VAR_GLOBAL   // PLC tag table "Carrier_SDC_TagTable"
   "Carrier_01_Status" AT %IW400 : Word;   // CARRIER STATUS WORD
   "Carrier_01_Status.0" AT %I400.0 : Bool;   // HEARTBEAT
   "Carrier_01_Status.1" AT %I400.1 : Bool;   // MANUAL
   "Carrier_01_Status.2" AT %I400.2 : Bool;   // IN_AUTO
   "Carrier_01_Status.3" AT %I400.3 : Bool;   // POSITIONING_COMPLETE
   "Carrier_01_Status.4" AT %I400.4 : Bool;   // PRODUCTION HOLD
   "Carrier_01_Status.5" AT %I400.5 : Bool;   // CARRIER MOVING FORWARD
   "Carrier_01_Status.6" AT %I400.6 : Bool;   // CARRIER MOVING REVERSE
   "Carrier_01_Status.7" AT %I400.7 : Bool;   // CARRIER FAULT
   "Carrier_01_Status.8" AT %I401.0 : Bool;   // CRASH DETECT TRIPPED
   "Carrier_01_Status.9" AT %I401.1 : Bool;
   "Carrier_01_Status.10" AT %I401.2 : Bool;
   "Carrier_01_Status.11" AT %I401.3 : Bool;
   "Carrier_01_Status.12" AT %I401.4 : Bool;
   "Carrier_01_Status.13" AT %I401.5 : Bool;
   "Carrier_01_Status.14" AT %I401.6 : Bool;
   "Carrier_01_Status.15" AT %I401.7 : Bool;
   "Carrier_01_SDCFaultCode" AT %IW402 : Word;   // SDC FAULT CODE
   "Carrier_01_CarrierPosition" AT %ID404 : DWord;   // CARRIER POSITION
   "Carrier_01_CarrierNumber" AT %IW408 : Word;   // CARRIER NUMBER
   "Carrier_01_G120DControlWord" AT %IW410 : Word;   // G120D_STW1_CONTROL
   "Carrier_01_G120DControlWord.0" AT %I410.0 : Bool;   // Bit_00_ON
   "Carrier_01_G120DControlWord.1" AT %I410.1 : Bool;   // Bit_01_AUS2_INH
   "Carrier_01_G120DControlWord.2" AT %I410.2 : Bool;   // Bit_02_AUS3_STOP
   "Carrier_01_G120DControlWord.3" AT %I410.3 : Bool;   // Bit_03_EN
   "Carrier_01_G120DControlWord.4" AT %I410.4 : Bool;   // Bit_04_EN_RAMP
   "Carrier_01_G120DControlWord.5" AT %I410.5 : Bool;   // Bit_05_START_RAMP
   "Carrier_01_G120DControlWord.6" AT %I410.6 : Bool;   // Bit_06_SETPOINT
   "Carrier_01_G120DControlWord.7" AT %I410.7 : Bool;   // Bit_07_RESET
   "Carrier_01_G120DControlWord.8" AT %I411.0 : Bool;   // Bit_08_JOG_R
   "Carrier_01_G120DControlWord.9" AT %I411.1 : Bool;   // Bit_09_JOG_L
   "Carrier_01_G120DControlWord.10" AT %I411.2 : Bool;   // Bit_10_CONTR_PLC
   "Carrier_01_G120DControlWord.11" AT %I411.3 : Bool;   // Bit_11_REVERSE
   "Carrier_01_G120DControlWord.12" AT %I411.4 : Bool;   // Bit_12_BRAKE_RELEASE
   "Carrier_01_G120DControlWord.13" AT %I411.5 : Bool;   // Bit_13_DDS
   "Carrier_01_G120DControlWord.14" AT %I411.6 : Bool;   // Bit_14_DO0
   "Carrier_01_G120DControlWord.15" AT %I411.7 : Bool;   // Bit_15_DO1
   "Carrier_01_G120DStatusWord" AT %IW412 : Word;   // G120D_ZSW1_STATUS
   "Carrier_01_G120DStatusWord.0" AT %I412.0 : Bool;   // Bit_00_READY_RUN
   "Carrier_01_G120DStatusWord.1" AT %I412.1 : Bool;   // Bit_01_READY_ON
   "Carrier_01_G120DStatusWord.2" AT %I412.2 : Bool;   // Bit_02_ENABLE
   "Carrier_01_G120DStatusWord.3" AT %I412.3 : Bool;   // Bit_03_FAULT
   "Carrier_01_G120DStatusWord.4" AT %I412.4 : Bool;   // Bit_04_OFF2
   "Carrier_01_G120DStatusWord.5" AT %I412.5 : Bool;   // Bit_05_OFF3
   "Carrier_01_G120DStatusWord.6" AT %I412.6 : Bool;   // Bit_06_LOCK_OUT
   "Carrier_01_G120DStatusWord.7" AT %I412.7 : Bool;   // Bit_07_WARN
   "Carrier_01_G120DStatusWord.8" AT %I413.0 : Bool;   // Bit_08_NO_DEVIATION
   "Carrier_01_G120DStatusWord.9" AT %I413.1 : Bool;   // Bit_09_CONTR_PLC
   "Carrier_01_G120DStatusWord.10" AT %I413.2 : Bool;   // Bit_10_F_MAX
   "Carrier_01_G120DStatusWord.11" AT %I413.3 : Bool;   // Bit_11_LIMIT_REACHED
   "Carrier_01_G120DStatusWord.12" AT %I413.4 : Bool;   // Bit_12_BRAKE_OPEN
   "Carrier_01_G120DStatusWord.13" AT %I413.5 : Bool;   // Bit_13_NO_OVERTEMP
   "Carrier_01_G120DStatusWord.14" AT %I413.6 : Bool;   // Bit_14_CW_CCW
   "Carrier_01_G120DStatusWord.15" AT %I413.7 : Bool;   // Bit_15_OVERL
   "Carrier_01_Slot2_Input" AT %IW414 : Word;   // SLOT 2 INPUT WORD
   "Carrier_01_CrashDetectSW" AT %I414.0 : Bool;   // CRASH DETECT SW
   "Carrier_01_SpareSafetyInput(2_1)" AT %I414.1 : Bool;   // SPARE SAFETY INPUT
   "Carrier_01_SpareSafetyInput(2_2)" AT %I414.2 : Bool;   // SPARE SAFETY INPUT
   "Carrier_01_SpareSafetyInput(2_3)" AT %I414.3 : Bool;   // SPARE SAFETY INPUT
   "Carrier_01_SpareSafetyInput(2_4)" AT %I414.4 : Bool;   // SPARE SAFETY INPUT
   "Carrier_01_SpareSafetyInput(2_5)" AT %I414.5 : Bool;   // SPARE SAFETY INPUT
   "Carrier_01_SpareSafetyInput(2_6)" AT %I414.6 : Bool;   // SPARE SAFETY INPUT
   "Carrier_01_SpareSafetyInput(2_7)" AT %I414.7 : Bool;   // SPARE SAFETY INPUT
   "Carrier_01_Slot3_SafetyOutput" AT %IW415 : Word;   // SLOT 3 SAFETY OUTPUT WORD
   "Carrier_01_Crash_Detect_OK" AT %I415.0 : Bool;   // CARRIER CRASH DETECT
   "Carrier_01_SpareSafetyOutput(3_1)" AT %I415.1 : Bool;   // SPARE SAFETY OUTPUT
   "Carrier_01_SpareSafetyOutput(3_2)" AT %I415.2 : Bool;   // SPARE SAFETY OUTPUT
   "Carrier_01_SpareSafetyOutput(3_3)" AT %I415.3 : Bool;   // SPARE SAFETY OUTPUT
   "Carrier_01_SpareSafetyOutput(3_4)" AT %I415.4 : Bool;   // SPARE SAFETY OUTPUT
   "Carrier_01_SpareSafetyOutput(3_5)" AT %I415.5 : Bool;   // SPARE SAFETY OUTPUT
   "Carrier_01_SpareSafetyOutput(3_6)" AT %I415.6 : Bool;   // SPARE SAFETY OUTPUT
   "Carrier_01_SpareSafetyOutput(3_7)" AT %I415.7 : Bool;   // SPARE SAFETY OUTPUT
   "Carrier_01_Slot4_Input" AT %IW416 : Word;   // SLOT 4 INPUT WORD
   "Carrier_01_480VPowerOn_MDCB1" AT %I416.0 : Bool;   // 480 VAC POWER ON MDCB 1
   "Carrier_01_SpareInput(4_1)" AT %I416.1 : Bool;   // SPARE INPUT
   "Carrier_01_SpareInput(4_2)" AT %I416.2 : Bool;   // SPARE INPUT
   "Carrier_01_SitopSelectStatus" AT %I416.3 : Bool;   // SITOP SELECT STATUS
   "Carrier_01_DCsupplyOnPSCB2" AT %I416.4 : Bool;   // DC SUPPLY ON PSCB 2
   "Carrier_01_SpareInput(4_5)" AT %I416.5 : Bool;   // SPARE INPUT
   "Carrier_01_SpareInput(4_6)" AT %I416.6 : Bool;   // SPARE INPUT
   "Carrier_01_SpareInput(4_7)" AT %I416.7 : Bool;   // SPARE INPUT
   "Carrier_01_PB1_ProdHoldLH" AT %I417.0 : Bool;   // PB 1 PRODUCTION HOLD LH
   "Carrier_01_PB2_ResetLH" AT %I417.1 : Bool;   // PB 2 RESET LH
   "Carrier_01_PB3_ProdHoldRH" AT %I417.2 : Bool;   // PB 3 PRODUCTION HOLD RH
   "Carrier_01_PB4_ResetRH" AT %I417.3 : Bool;   // PB 4 RESET RH
   "Carrier_01_SpareInput(4_14)" AT %I417.4 : Bool;   // SPARE INPUT
   "Carrier_01_SpareInput(4_15)" AT %I417.5 : Bool;   // SPARE INPUT
   "Carrier_01_SpareInput(4_16)" AT %I417.6 : Bool;   // SPARE INPUT
   "Carrier_01_SpareInput(4_17)" AT %I417.7 : Bool;   // SPARE INPUT
   "Carrier_01_Slot5_Output" AT %IW418 : Word;   // SLOT 5 OUTPUT WORD
   "Carrier_01_IRD400_HMI_24VDC_ENABLE" AT %I418.0 : Bool;   // IRD 400 PANEL HMI 24V DC POWER
   "Carrier_01_FaultLight_LH" AT %I418.1 : Bool;   // FAULT LIGHT LH
   "Carrier_01_RunLight_LH" AT %I418.2 : Bool;   // RUN LIGHT LH
   "Carrier_01_FaultLight_RH" AT %I418.3 : Bool;   // FAULT LIGHT RH
   "Carrier_01_RunLight_RH" AT %I418.4 : Bool;   // RUN LIGHT RH
   "Carrier_01_SpareOutput(5_5)" AT %I418.5 : Bool;   // SPARE OUTPUT
   "Carrier_01_SpareOutput(5_6)" AT %I418.6 : Bool;   // SPARE OUTPUT
   "Carrier_01_SpareOutput(5_7)" AT %I418.7 : Bool;   // SPARE OUTPUT
   "Carrier_01_ActualSpeed" AT %IW420 : Word;   // ACTUAL SPEED
   "Carrier_01_CarrierDriveAlarm" AT %IW422 : Word;   // CARRIER DRIVE ALARM
   "Carrier_01_CarrierDriveWarning" AT %IW424 : Word;   // CARRIER DRIVE WARNING
   "Carrier_02_Status" AT %IW450 : Word;   // CARRIER STATUS WORD
   "Carrier_02_Status.0" AT %I450.0 : Bool;   // HEARTBEAT
   "Carrier_02_Status.1" AT %I450.1 : Bool;   // MANUAL
   "Carrier_02_Status.2" AT %I450.2 : Bool;   // IN_AUTO
   "Carrier_02_Status.3" AT %I450.3 : Bool;   // POSITIONING_COMPLETE
   "Carrier_02_Status.4" AT %I450.4 : Bool;   // PRODUCTION HOLD
   "Carrier_02_Status.5" AT %I450.5 : Bool;   // CARRIER MOVING FORWARD
   "Carrier_02_Status.6" AT %I450.6 : Bool;   // CARRIER MOVING REVERSE
   "Carrier_02_Status.7" AT %I450.7 : Bool;   // CARRIER FAULT
   "Carrier_02_Status.8" AT %I451.0 : Bool;   // CRASH DETECT TRIPPED
   "Carrier_02_Status.9" AT %I451.1 : Bool;
   "Carrier_02_Status.10" AT %I451.2 : Bool;
   "Carrier_02_Status.11" AT %I451.3 : Bool;
   "Carrier_02_Status.12" AT %I451.4 : Bool;
   "Carrier_02_Status.13" AT %I451.5 : Bool;
   "Carrier_02_Status.14" AT %I451.6 : Bool;
   "Carrier_02_Status.15" AT %I451.7 : Bool;
   "Carrier_02_SDCFaultCode" AT %IW452 : Word;   // SDC FAULT CODE
   "Carrier_02_CarrierPosition" AT %ID454 : DWord;   // CARRIER POSITION
   "Carrier_02_CarrierNumber" AT %IW458 : Word;   // CARRIER NUMBER
   "Carrier_02_G120DControlWord" AT %IW460 : Word;   // G120D_STW1_CONTROL
   "Carrier_02_G120DControlWord.0" AT %I460.0 : Bool;   // Bit_00_ON
   "Carrier_02_G120DControlWord.1" AT %I460.1 : Bool;   // Bit_01_AUS2_INH
   "Carrier_02_G120DControlWord.2" AT %I460.2 : Bool;   // Bit_02_AUS3_STOP
   "Carrier_02_G120DControlWord.3" AT %I460.3 : Bool;   // Bit_03_EN
   "Carrier_02_G120DControlWord.4" AT %I460.4 : Bool;   // Bit_04_EN_RAMP
   "Carrier_02_G120DControlWord.5" AT %I460.5 : Bool;   // Bit_05_START_RAMP
   "Carrier_02_G120DControlWord.6" AT %I460.6 : Bool;   // Bit_06_SETPOINT
   "Carrier_02_G120DControlWord.7" AT %I460.7 : Bool;   // Bit_07_RESET
   "Carrier_02_G120DControlWord.8" AT %I461.0 : Bool;   // Bit_08_JOG_R
   "Carrier_02_G120DControlWord.9" AT %I461.1 : Bool;   // Bit_09_JOG_L
   "Carrier_02_G120DControlWord.10" AT %I461.2 : Bool;   // Bit_10_CONTR_PLC
   "Carrier_02_G120DControlWord.11" AT %I461.3 : Bool;   // Bit_11_REVERSE
   "Carrier_02_G120DControlWord.12" AT %I461.4 : Bool;   // Bit_12_BRAKE_RELEASE
   "Carrier_02_G120DControlWord.13" AT %I461.5 : Bool;   // Bit_13_DDS
   "Carrier_02_G120DControlWord.14" AT %I461.6 : Bool;   // Bit_14_DO0
   "Carrier_02_G120DControlWord.15" AT %I461.7 : Bool;   // Bit_15_DO1
   "Carrier_02_G120DStatusWord" AT %IW462 : Word;   // G120D_ZSW1_STATUS
   "Carrier_02_G120DStatusWord.0" AT %I462.0 : Bool;   // Bit_00_READY_RUN
   "Carrier_02_G120DStatusWord.1" AT %I462.1 : Bool;   // Bit_01_READY_ON
   "Carrier_02_G120DStatusWord.2" AT %I462.2 : Bool;   // Bit_02_ENABLE
   "Carrier_02_G120DStatusWord.3" AT %I462.3 : Bool;   // Bit_03_FAULT
   "Carrier_02_G120DStatusWord.4" AT %I462.4 : Bool;   // Bit_04_OFF2
   "Carrier_02_G120DStatusWord.5" AT %I462.5 : Bool;   // Bit_05_OFF3
   "Carrier_02_G120DStatusWord.6" AT %I462.6 : Bool;   // Bit_06_LOCK_OUT
   "Carrier_02_G120DStatusWord.7" AT %I462.7 : Bool;   // Bit_07_WARN
   "Carrier_02_G120DStatusWord.8" AT %I463.0 : Bool;   // Bit_08_NO_DEVIATION
   "Carrier_02_G120DStatusWord.9" AT %I463.1 : Bool;   // Bit_09_CONTR_PLC
   "Carrier_02_G120DStatusWord.10" AT %I463.2 : Bool;   // Bit_10_F_MAX
   "Carrier_02_G120DStatusWord.11" AT %I463.3 : Bool;   // Bit_11_LIMIT_REACHED
   "Carrier_02_G120DStatusWord.12" AT %I463.4 : Bool;   // Bit_12_BRAKE_OPEN
   "Carrier_02_G120DStatusWord.13" AT %I463.5 : Bool;   // Bit_13_NO_OVERTEMP
   "Carrier_02_G120DStatusWord.14" AT %I463.6 : Bool;   // Bit_14_CW_CCW
   "Carrier_02_G120DStatusWord.15" AT %I463.7 : Bool;   // Bit_15_OVERL
   "Carrier_02_Slot2_Input" AT %IW464 : Word;   // SLOT 2 INPUT WORD
   "Carrier_02_CrashDetectSW" AT %I464.0 : Bool;   // CRASH DETECT SW
   "Carrier_02_SpareSafetyInput(2_1)" AT %I464.1 : Bool;   // SPARE SAFETY INPUT
   "Carrier_02_SpareSafetyInput(2_2)" AT %I464.2 : Bool;   // SPARE SAFETY INPUT
   "Carrier_02_SpareSafetyInput(2_3)" AT %I464.3 : Bool;   // SPARE SAFETY INPUT
   "Carrier_02_SpareSafetyInput(2_4)" AT %I464.4 : Bool;   // SPARE SAFETY INPUT
   "Carrier_02_SpareSafetyInput(2_5)" AT %I464.5 : Bool;   // SPARE SAFETY INPUT
   "Carrier_02_SpareSafetyInput(2_6)" AT %I464.6 : Bool;   // SPARE SAFETY INPUT
   "Carrier_02_SpareSafetyInput(2_7)" AT %I464.7 : Bool;   // SPARE SAFETY INPUT
   "Carrier_02_Slot3_SafetyOutput" AT %IW465 : Word;   // SLOT 3 SAFETY OUTPUT WORD
   "Carrier_02_Crash_Detect_OK" AT %I465.0 : Bool;   // CARRIER CRASH DETECT
   "Carrier_02_SpareSafetyOutput(3_1)" AT %I465.1 : Bool;   // SPARE SAFETY OUTPUT
   "Carrier_02_SpareSafetyOutput(3_2)" AT %I465.2 : Bool;   // SPARE SAFETY OUTPUT
   "Carrier_02_SpareSafetyOutput(3_3)" AT %I465.3 : Bool;   // SPARE SAFETY OUTPUT
   "Carrier_02_SpareSafetyOutput(3_4)" AT %I465.4 : Bool;   // SPARE SAFETY OUTPUT
   "Carrier_02_SpareSafetyOutput(3_5)" AT %I465.5 : Bool;   // SPARE SAFETY OUTPUT
   "Carrier_02_SpareSafetyOutput(3_6)" AT %I465.6 : Bool;   // SPARE SAFETY OUTPUT
   "Carrier_02_SpareSafetyOutput(3_7)" AT %I465.7 : Bool;   // SPARE SAFETY OUTPUT
   "Carrier_02_Slot4_Input" AT %IW466 : Word;   // SLOT 4 INPUT WORD
   "Carrier_02_480VPowerOn_MDCB1" AT %I466.0 : Bool;   // 480 VAC POWER ON MDCB 1
   "Carrier_02_SpareInput(4_1)" AT %I466.1 : Bool;   // SPARE INPUT
   "Carrier_02_SpareInput(4_2)" AT %I466.2 : Bool;   // SPARE INPUT
   "Carrier_02_SitopSelectStatus" AT %I466.3 : Bool;   // SITOP SELECT STATUS
   "Carrier_02_DCsupplyOnPSCB2" AT %I466.4 : Bool;   // DC SUPPLY ON PSCB 2
   "Carrier_02_SpareInput(4_5)" AT %I466.5 : Bool;   // SPARE INPUT
   "Carrier_02_SpareInput(4_6)" AT %I466.6 : Bool;   // SPARE INPUT
   "Carrier_02_SpareInput(4_7)" AT %I466.7 : Bool;   // SPARE INPUT
   "Carrier_02_PB1_ProdHoldLH" AT %I467.0 : Bool;   // PB 1 PRODUCTION HOLD LH
   "Carrier_02_PB2_ResetLH" AT %I467.1 : Bool;   // PB 2 RESET LH
   "Carrier_02_PB3_ProdHoldRH" AT %I467.2 : Bool;   // PB 3 PRODUCTION HOLD RH
   "Carrier_02_PB4_ResetRH" AT %I467.3 : Bool;   // PB 4 RESET RH
   "Carrier_02_SpareInput(4_14)" AT %I467.4 : Bool;   // SPARE INPUT
   "Carrier_02_SpareInput(4_15)" AT %I467.5 : Bool;   // SPARE INPUT
   "Carrier_02_SpareInput(4_16)" AT %I467.6 : Bool;   // SPARE INPUT
   "Carrier_02_SpareInput(4_17)" AT %I467.7 : Bool;   // SPARE INPUT
   "Carrier_02_Slot5_Output" AT %IW468 : Word;   // SLOT 5 OUTPUT WORD
   "Carrier_02_IRD400_HMI_24VDC_ENABLE" AT %I468.0 : Bool;   // IRD 400 PANEL HMI 24V DC POWER
   "Carrier_02_FaultLight_LH" AT %I468.1 : Bool;   // FAULT LIGHT LH
   "Carrier_02_RunLight_LH" AT %I468.2 : Bool;   // RUN LIGHT LH
   "Carrier_02_FaultLight_RH" AT %I468.3 : Bool;   // FAULT LIGHT RH
   "Carrier_02_RunLight_RH" AT %I468.4 : Bool;   // RUN LIGHT RH
   "Carrier_02_SpareOutput(5_5)" AT %I468.5 : Bool;   // SPARE OUTPUT
   "Carrier_02_SpareOutput(5_6)" AT %I468.6 : Bool;   // SPARE OUTPUT
   "Carrier_02_SpareOutput(5_7)" AT %I468.7 : Bool;   // SPARE OUTPUT
   "Carrier_02_ActualSpeed" AT %IW470 : Word;   // ACTUAL SPEED
   "Carrier_02_CarrierDriveAlarm" AT %IW472 : Word;   // CARRIER DRIVE ALARM
   "Carrier_02_CarrierDriveWarning" AT %IW474 : Word;   // CARRIER DRIVE WARNING
   "Carrier_03_Status" AT %IW500 : Word;   // CARRIER STATUS WORD
   "Carrier_03_Status.0" AT %I500.0 : Bool;   // HEARTBEAT
   "Carrier_03_Status.1" AT %I500.1 : Bool;   // MANUAL
   "Carrier_03_Status.2" AT %I500.2 : Bool;   // IN_AUTO
   "Carrier_03_Status.3" AT %I500.3 : Bool;   // POSITIONING_COMPLETE
   "Carrier_03_Status.4" AT %I500.4 : Bool;   // PRODUCTION HOLD
   "Carrier_03_Status.5" AT %I500.5 : Bool;   // CARRIER MOVING FORWARD
   "Carrier_03_Status.6" AT %I500.6 : Bool;   // CARRIER MOVING REVERSE
   "Carrier_03_Status.7" AT %I500.7 : Bool;   // CARRIER FAULT
   "Carrier_03_Status.8" AT %I501.0 : Bool;   // CRASH DETECT TRIPPED
   "Carrier_03_Status.9" AT %I501.1 : Bool;
   "Carrier_03_Status.10" AT %I501.2 : Bool;
   "Carrier_03_Status.11" AT %I501.3 : Bool;
   "Carrier_03_Status.12" AT %I501.4 : Bool;
   "Carrier_03_Status.13" AT %I501.5 : Bool;
   "Carrier_03_Status.14" AT %I501.6 : Bool;
   "Carrier_03_Status.15" AT %I501.7 : Bool;
   "Carrier_03_SDCFaultCode" AT %IW502 : Word;   // SDC FAULT CODE
   "Carrier_03_CarrierPosition" AT %ID504 : DWord;   // CARRIER POSITION
   "Carrier_03_CarrierNumber" AT %IW508 : Word;   // CARRIER NUMBER
   "Carrier_03_G120DControlWord" AT %IW510 : Word;   // G120D_STW1_CONTROL
   "Carrier_03_G120DControlWord.0" AT %I510.0 : Bool;   // Bit_00_ON
   "Carrier_03_G120DControlWord.1" AT %I510.1 : Bool;   // Bit_01_AUS2_INH
   "Carrier_03_G120DControlWord.2" AT %I510.2 : Bool;   // Bit_02_AUS3_STOP
   "Carrier_03_G120DControlWord.3" AT %I510.3 : Bool;   // Bit_03_EN
   "Carrier_03_G120DControlWord.4" AT %I510.4 : Bool;   // Bit_04_EN_RAMP
   "Carrier_03_G120DControlWord.5" AT %I510.5 : Bool;   // Bit_05_START_RAMP
   "Carrier_03_G120DControlWord.6" AT %I510.6 : Bool;   // Bit_06_SETPOINT
   "Carrier_03_G120DControlWord.7" AT %I510.7 : Bool;   // Bit_07_RESET
   "Carrier_03_G120DControlWord.8" AT %I511.0 : Bool;   // Bit_08_JOG_R
   "Carrier_03_G120DControlWord.9" AT %I511.1 : Bool;   // Bit_09_JOG_L
   "Carrier_03_G120DControlWord.10" AT %I511.2 : Bool;   // Bit_10_CONTR_PLC
   "Carrier_03_G120DControlWord.11" AT %I511.3 : Bool;   // Bit_11_REVERSE
   "Carrier_03_G120DControlWord.12" AT %I511.4 : Bool;   // Bit_12_BRAKE_RELEASE
   "Carrier_03_G120DControlWord.13" AT %I511.5 : Bool;   // Bit_13_DDS
   "Carrier_03_G120DControlWord.14" AT %I511.6 : Bool;   // Bit_14_DO0
   "Carrier_03_G120DControlWord.15" AT %I511.7 : Bool;   // Bit_15_DO1
   "Carrier_03_G120DStatusWord" AT %IW512 : Word;   // G120D_ZSW1_STATUS
   "Carrier_03_G120DStatusWord.0" AT %I512.0 : Bool;   // Bit_00_READY_RUN
   "Carrier_03_G120DStatusWord.1" AT %I512.1 : Bool;   // Bit_01_READY_ON
   "Carrier_03_G120DStatusWord.2" AT %I512.2 : Bool;   // Bit_02_ENABLE
   "Carrier_03_G120DStatusWord.3" AT %I512.3 : Bool;   // Bit_03_FAULT
   "Carrier_03_G120DStatusWord.4" AT %I512.4 : Bool;   // Bit_04_OFF2
   "Carrier_03_G120DStatusWord.5" AT %I512.5 : Bool;   // Bit_05_OFF3
   "Carrier_03_G120DStatusWord.6" AT %I512.6 : Bool;   // Bit_06_LOCK_OUT
   "Carrier_03_G120DStatusWord.7" AT %I512.7 : Bool;   // Bit_07_WARN
   "Carrier_03_G120DStatusWord.8" AT %I513.0 : Bool;   // Bit_08_NO_DEVIATION
   "Carrier_03_G120DStatusWord.9" AT %I513.1 : Bool;   // Bit_09_CONTR_PLC
   "Carrier_03_G120DStatusWord.10" AT %I513.2 : Bool;   // Bit_10_F_MAX
   "Carrier_03_G120DStatusWord.11" AT %I513.3 : Bool;   // Bit_11_LIMIT_REACHED
   "Carrier_03_G120DStatusWord.12" AT %I513.4 : Bool;   // Bit_12_BRAKE_OPEN
   "Carrier_03_G120DStatusWord.13" AT %I513.5 : Bool;   // Bit_13_NO_OVERTEMP
   "Carrier_03_G120DStatusWord.14" AT %I513.6 : Bool;   // Bit_14_CW_CCW
   "Carrier_03_G120DStatusWord.15" AT %I513.7 : Bool;   // Bit_15_OVERL
   "Carrier_03_Slot2_Input" AT %IW514 : Word;   // SLOT 2 INPUT WORD
   "Carrier_03_CrashDetectSW" AT %I514.0 : Bool;   // CRASH DETECT SW
   "Carrier_03_SpareSafetyInput(2_1)" AT %I514.1 : Bool;   // SPARE SAFETY INPUT
   "Carrier_03_SpareSafetyInput(2_2)" AT %I514.2 : Bool;   // SPARE SAFETY INPUT
   "Carrier_03_SpareSafetyInput(2_3)" AT %I514.3 : Bool;   // SPARE SAFETY INPUT
   "Carrier_03_SpareSafetyInput(2_4)" AT %I514.4 : Bool;   // SPARE SAFETY INPUT
   "Carrier_03_SpareSafetyInput(2_5)" AT %I514.5 : Bool;   // SPARE SAFETY INPUT
   "Carrier_03_SpareSafetyInput(2_6)" AT %I514.6 : Bool;   // SPARE SAFETY INPUT
   "Carrier_03_SpareSafetyInput(2_7)" AT %I514.7 : Bool;   // SPARE SAFETY INPUT
   "Carrier_03_Slot3_SafetyOutput" AT %IW515 : Word;   // SLOT 3 SAFETY OUTPUT WORD
   "Carrier_03_Crash_Detect_OK" AT %I515.0 : Bool;   // CARRIER CRASH DETECT
   "Carrier_03_SpareSafetyOutput(3_1)" AT %I515.1 : Bool;   // SPARE SAFETY OUTPUT
   "Carrier_03_SpareSafetyOutput(3_2)" AT %I515.2 : Bool;   // SPARE SAFETY OUTPUT
   "Carrier_03_SpareSafetyOutput(3_3)" AT %I515.3 : Bool;   // SPARE SAFETY OUTPUT
   "Carrier_03_SpareSafetyOutput(3_4)" AT %I515.4 : Bool;   // SPARE SAFETY OUTPUT
   "Carrier_03_SpareSafetyOutput(3_5)" AT %I515.5 : Bool;   // SPARE SAFETY OUTPUT
   "Carrier_03_SpareSafetyOutput(3_6)" AT %I515.6 : Bool;   // SPARE SAFETY OUTPUT
   "Carrier_03_SpareSafetyOutput(3_7)" AT %I515.7 : Bool;   // SPARE SAFETY OUTPUT
   "Carrier_03_Slot4_Input" AT %IW516 : Word;   // SLOT 4 INPUT WORD
   "Carrier_03_480VPowerOn_MDCB1" AT %I516.0 : Bool;   // 480 VAC POWER ON MDCB 1
   "Carrier_03_SpareInput(4_1)" AT %I516.1 : Bool;   // SPARE INPUT
   "Carrier_03_SpareInput(4_2)" AT %I516.2 : Bool;   // SPARE INPUT
   "Carrier_03_SitopSelectStatus" AT %I516.3 : Bool;   // SITOP SELECT STATUS
   "Carrier_03_DCsupplyOnPSCB2" AT %I516.4 : Bool;   // DC SUPPLY ON PSCB 2
   "Carrier_03_SpareInput(4_5)" AT %I516.5 : Bool;   // SPARE INPUT
   "Carrier_03_SpareInput(4_6)" AT %I516.6 : Bool;   // SPARE INPUT
   "Carrier_03_SpareInput(4_7)" AT %I516.7 : Bool;   // SPARE INPUT
   "Carrier_03_PB1_ProdHoldLH" AT %I517.0 : Bool;   // PB 1 PRODUCTION HOLD LH
   "Carrier_03_PB2_ResetLH" AT %I517.1 : Bool;   // PB 2 RESET LH
   "Carrier_03_PB3_ProdHoldRH" AT %I517.2 : Bool;   // PB 3 PRODUCTION HOLD RH
   "Carrier_03_PB4_ResetRH" AT %I517.3 : Bool;   // PB 4 RESET RH
   "Carrier_03_SpareInput(4_14)" AT %I517.4 : Bool;   // SPARE INPUT
   "Carrier_03_SpareInput(4_15)" AT %I517.5 : Bool;   // SPARE INPUT
   "Carrier_03_SpareInput(4_16)" AT %I517.6 : Bool;   // SPARE INPUT
   "Carrier_03_SpareInput(4_17)" AT %I517.7 : Bool;   // SPARE INPUT
   "Carrier_03_Slot5_Output" AT %IW518 : Word;   // SLOT 5 OUTPUT WORD
   "Carrier_03_IRD400_HMI_24VDC_ENABLE" AT %I518.0 : Bool;   // IRD 400 PANEL HMI 24V DC POWER
   "Carrier_03_FaultLight_LH" AT %I518.1 : Bool;   // FAULT LIGHT LH
   "Carrier_03_RunLight_LH" AT %I518.2 : Bool;   // RUN LIGHT LH
   "Carrier_03_FaultLight_RH" AT %I518.3 : Bool;   // FAULT LIGHT RH
   "Carrier_03_RunLight_RH" AT %I518.4 : Bool;   // RUN LIGHT RH
   "Carrier_03_SpareOutput(5_5)" AT %I518.5 : Bool;   // SPARE OUTPUT
   "Carrier_03_SpareOutput(5_6)" AT %I518.6 : Bool;   // SPARE OUTPUT
   "Carrier_03_SpareOutput(5_7)" AT %I518.7 : Bool;   // SPARE OUTPUT
   "Carrier_03_ActualSpeed" AT %IW520 : Word;   // ACTUAL SPEED
   "Carrier_03_CarrierDriveAlarm" AT %IW522 : Word;   // CARRIER DRIVE ALARM
   "Carrier_03_CarrierDriveWarning" AT %IW524 : Word;   // CARRIER DRIVE WARNING
   "Carrier_04_Status" AT %IW550 : Word;   // CARRIER STATUS WORD
   "Carrier_04_Status.0" AT %I550.0 : Bool;   // HEARTBEAT
   "Carrier_04_Status.1" AT %I550.1 : Bool;   // MANUAL
   "Carrier_04_Status.2" AT %I550.2 : Bool;   // IN_AUTO
   "Carrier_04_Status.3" AT %I550.3 : Bool;   // POSITIONING_COMPLETE
   "Carrier_04_Status.4" AT %I550.4 : Bool;   // PRODUCTION HOLD
   "Carrier_04_Status.5" AT %I550.5 : Bool;   // CARRIER MOVING FORWARD
   "Carrier_04_Status.6" AT %I550.6 : Bool;   // CARRIER MOVING REVERSE
   "Carrier_04_Status.7" AT %I550.7 : Bool;   // CARRIER FAULT
   "Carrier_04_Status.8" AT %I551.0 : Bool;   // CRASH DETECT TRIPPED
   "Carrier_04_Status.9" AT %I551.1 : Bool;
   "Carrier_04_Status.10" AT %I551.2 : Bool;
   "Carrier_04_Status.11" AT %I551.3 : Bool;
   "Carrier_04_Status.12" AT %I551.4 : Bool;
   "Carrier_04_Status.13" AT %I551.5 : Bool;
   "Carrier_04_Status.14" AT %I551.6 : Bool;
   "Carrier_04_Status.15" AT %I551.7 : Bool;
   "Carrier_04_SDCFaultCode" AT %IW552 : Word;   // SDC FAULT CODE
   "Carrier_04_CarrierPosition" AT %ID554 : DWord;   // CARRIER POSITION
   "Carrier_04_CarrierNumber" AT %IW558 : Word;   // CARRIER NUMBER
   "Carrier_04_G120DControlWord" AT %IW560 : Word;   // G120D_STW1_CONTROL
   "Carrier_04_G120DControlWord.0" AT %I560.0 : Bool;   // Bit_00_ON
   "Carrier_04_G120DControlWord.1" AT %I560.1 : Bool;   // Bit_01_AUS2_INH
   "Carrier_04_G120DControlWord.2" AT %I560.2 : Bool;   // Bit_02_AUS3_STOP
   "Carrier_04_G120DControlWord.3" AT %I560.3 : Bool;   // Bit_03_EN
   "Carrier_04_G120DControlWord.4" AT %I560.4 : Bool;   // Bit_04_EN_RAMP
   "Carrier_04_G120DControlWord.5" AT %I560.5 : Bool;   // Bit_05_START_RAMP
   "Carrier_04_G120DControlWord.6" AT %I560.6 : Bool;   // Bit_06_SETPOINT
   "Carrier_04_G120DControlWord.7" AT %I560.7 : Bool;   // Bit_07_RESET
   "Carrier_04_G120DControlWord.8" AT %I561.0 : Bool;   // Bit_08_JOG_R
   "Carrier_04_G120DControlWord.9" AT %I561.1 : Bool;   // Bit_09_JOG_L
   "Carrier_04_G120DControlWord.10" AT %I561.2 : Bool;   // Bit_10_CONTR_PLC
   "Carrier_04_G120DControlWord.11" AT %I561.3 : Bool;   // Bit_11_REVERSE
   "Carrier_04_G120DControlWord.12" AT %I561.4 : Bool;   // Bit_12_BRAKE_RELEASE
   "Carrier_04_G120DControlWord.13" AT %I561.5 : Bool;   // Bit_13_DDS
   "Carrier_04_G120DControlWord.14" AT %I561.6 : Bool;   // Bit_14_DO0
   "Carrier_04_G120DControlWord.15" AT %I561.7 : Bool;   // Bit_15_DO1
   "Carrier_04_G120DStatusWord" AT %IW562 : Word;   // G120D_ZSW1_STATUS
   "Carrier_04_G120DStatusWord.0" AT %I562.0 : Bool;   // Bit_00_READY_RUN
   "Carrier_04_G120DStatusWord.1" AT %I562.1 : Bool;   // Bit_01_READY_ON
   "Carrier_04_G120DStatusWord.2" AT %I562.2 : Bool;   // Bit_02_ENABLE
   "Carrier_04_G120DStatusWord.3" AT %I562.3 : Bool;   // Bit_03_FAULT
   "Carrier_04_G120DStatusWord.4" AT %I562.4 : Bool;   // Bit_04_OFF2
   "Carrier_04_G120DStatusWord.5" AT %I562.5 : Bool;   // Bit_05_OFF3
   "Carrier_04_G120DStatusWord.6" AT %I562.6 : Bool;   // Bit_06_LOCK_OUT
   "Carrier_04_G120DStatusWord.7" AT %I562.7 : Bool;   // Bit_07_WARN
   "Carrier_04_G120DStatusWord.8" AT %I563.0 : Bool;   // Bit_08_NO_DEVIATION
   "Carrier_04_G120DStatusWord.9" AT %I563.1 : Bool;   // Bit_09_CONTR_PLC
   "Carrier_04_G120DStatusWord.10" AT %I563.2 : Bool;   // Bit_10_F_MAX
   "Carrier_04_G120DStatusWord.11" AT %I563.3 : Bool;   // Bit_11_LIMIT_REACHED
   "Carrier_04_G120DStatusWord.12" AT %I563.4 : Bool;   // Bit_12_BRAKE_OPEN
   "Carrier_04_G120DStatusWord.13" AT %I563.5 : Bool;   // Bit_13_NO_OVERTEMP
   "Carrier_04_G120DStatusWord.14" AT %I563.6 : Bool;   // Bit_14_CW_CCW
   "Carrier_04_G120DStatusWord.15" AT %I563.7 : Bool;   // Bit_15_OVERL
   "Carrier_04_Slot2_Input" AT %IW564 : Word;   // SLOT 2 INPUT WORD
   "Carrier_04_CrashDetectSW" AT %I564.0 : Bool;   // CRASH DETECT SW
   "Carrier_04_SpareSafetyInput(2_1)" AT %I564.1 : Bool;   // SPARE SAFETY INPUT
   "Carrier_04_SpareSafetyInput(2_2)" AT %I564.2 : Bool;   // SPARE SAFETY INPUT
   "Carrier_04_SpareSafetyInput(2_3)" AT %I564.3 : Bool;   // SPARE SAFETY INPUT
   "Carrier_04_SpareSafetyInput(2_4)" AT %I564.4 : Bool;   // SPARE SAFETY INPUT
   "Carrier_04_SpareSafetyInput(2_5)" AT %I564.5 : Bool;   // SPARE SAFETY INPUT
   "Carrier_04_SpareSafetyInput(2_6)" AT %I564.6 : Bool;   // SPARE SAFETY INPUT
   "Carrier_04_SpareSafetyInput(2_7)" AT %I564.7 : Bool;   // SPARE SAFETY INPUT
   "Carrier_04_Slot3_SafetyOutput" AT %IW565 : Word;   // SLOT 3 SAFETY OUTPUT WORD
   "Carrier_04_Crash_Detect_OK" AT %I565.0 : Bool;   // CARRIER CRASH DETECT
   "Carrier_04_SpareSafetyOutput(3_1)" AT %I565.1 : Bool;   // SPARE SAFETY OUTPUT
   "Carrier_04_SpareSafetyOutput(3_2)" AT %I565.2 : Bool;   // SPARE SAFETY OUTPUT
   "Carrier_04_SpareSafetyOutput(3_3)" AT %I565.3 : Bool;   // SPARE SAFETY OUTPUT
   "Carrier_04_SpareSafetyOutput(3_4)" AT %I565.4 : Bool;   // SPARE SAFETY OUTPUT
   "Carrier_04_SpareSafetyOutput(3_5)" AT %I565.5 : Bool;   // SPARE SAFETY OUTPUT
   "Carrier_04_SpareSafetyOutput(3_6)" AT %I565.6 : Bool;   // SPARE SAFETY OUTPUT
   "Carrier_04_SpareSafetyOutput(3_7)" AT %I565.7 : Bool;   // SPARE SAFETY OUTPUT
   "Carrier_04_Slot4_Input" AT %IW566 : Word;   // SLOT 4 INPUT WORD
   "Carrier_04_480VPowerOn_MDCB1" AT %I566.0 : Bool;   // 480 VAC POWER ON MDCB 1
   "Carrier_04_SpareInput(4_1)" AT %I566.1 : Bool;   // SPARE INPUT
   "Carrier_04_SpareInput(4_2)" AT %I566.2 : Bool;   // SPARE INPUT
   "Carrier_04_SitopSelectStatus" AT %I566.3 : Bool;   // SITOP SELECT STATUS
   "Carrier_04_DCsupplyOnPSCB2" AT %I566.4 : Bool;   // DC SUPPLY ON PSCB 2
   "Carrier_04_SpareInput(4_5)" AT %I566.5 : Bool;   // SPARE INPUT
   "Carrier_04_SpareInput(4_6)" AT %I566.6 : Bool;   // SPARE INPUT
   "Carrier_04_SpareInput(4_7)" AT %I566.7 : Bool;   // SPARE INPUT
   "Carrier_04_PB1_ProdHoldLH" AT %I567.0 : Bool;   // PB 1 PRODUCTION HOLD LH
   "Carrier_04_PB2_ResetLH" AT %I567.1 : Bool;   // PB 2 RESET LH
   "Carrier_04_PB3_ProdHoldRH" AT %I567.2 : Bool;   // PB 3 PRODUCTION HOLD RH
   "Carrier_04_PB4_ResetRH" AT %I567.3 : Bool;   // PB 4 RESET RH
   "Carrier_04_SpareInput(4_14)" AT %I567.4 : Bool;   // SPARE INPUT
   "Carrier_04_SpareInput(4_15)" AT %I567.5 : Bool;   // SPARE INPUT
   "Carrier_04_SpareInput(4_16)" AT %I567.6 : Bool;   // SPARE INPUT
   "Carrier_04_SpareInput(4_17)" AT %I567.7 : Bool;   // SPARE INPUT
   "Carrier_04_Slot5_Output" AT %IW568 : Word;   // SLOT 5 OUTPUT WORD
   "Carrier_04_IRD400_HMI_24VDC_ENABLE" AT %I568.0 : Bool;   // IRD 400 PANEL HMI 24V DC POWER
   "Carrier_04_FaultLight_LH" AT %I568.1 : Bool;   // FAULT LIGHT LH
   "Carrier_04_RunLight_LH" AT %I568.2 : Bool;   // RUN LIGHT LH
   "Carrier_04_FaultLight_RH" AT %I568.3 : Bool;   // FAULT LIGHT RH
   "Carrier_04_RunLight_RH" AT %I568.4 : Bool;   // RUN LIGHT RH
   "Carrier_04_SpareOutput(5_5)" AT %I568.5 : Bool;   // SPARE OUTPUT
   "Carrier_04_SpareOutput(5_6)" AT %I568.6 : Bool;   // SPARE OUTPUT
   "Carrier_04_SpareOutput(5_7)" AT %I568.7 : Bool;   // SPARE OUTPUT
   "Carrier_04_ActualSpeed" AT %IW570 : Word;   // ACTUAL SPEED
   "Carrier_04_CarrierDriveAlarm" AT %IW572 : Word;   // CARRIER DRIVE ALARM
   "Carrier_04_CarrierDriveWarning" AT %IW574 : Word;   // CARRIER DRIVE WARNING
   "Carrier_05_Status" AT %IW600 : Word;   // CARRIER STATUS WORD
   "Carrier_05_Status.0" AT %I600.0 : Bool;   // HEARTBEAT
   "Carrier_05_Status.1" AT %I600.1 : Bool;   // MANUAL
   "Carrier_05_Status.2" AT %I600.2 : Bool;   // IN_AUTO
   "Carrier_05_Status.3" AT %I600.3 : Bool;   // POSITIONING_COMPLETE
   "Carrier_05_Status.4" AT %I600.4 : Bool;   // PRODUCTION HOLD
   "Carrier_05_Status.5" AT %I600.5 : Bool;   // CARRIER MOVING FORWARD
   "Carrier_05_Status.6" AT %I600.6 : Bool;   // CARRIER MOVING REVERSE
   "Carrier_05_Status.7" AT %I600.7 : Bool;   // CARRIER FAULT
   "Carrier_05_Status.8" AT %I601.0 : Bool;   // CRASH DETECT TRIPPED
   "Carrier_05_Status.9" AT %I601.1 : Bool;
   "Carrier_05_Status.10" AT %I601.2 : Bool;
   "Carrier_05_Status.11" AT %I601.3 : Bool;
   "Carrier_05_Status.12" AT %I601.4 : Bool;
   "Carrier_05_Status.13" AT %I601.5 : Bool;
   "Carrier_05_Status.14" AT %I601.6 : Bool;
   "Carrier_05_Status.15" AT %I601.7 : Bool;
   "Carrier_05_SDCFaultCode" AT %IW602 : Word;   // SDC FAULT CODE
   "Carrier_05_CarrierPosition" AT %ID604 : DWord;   // CARRIER POSITION
   "Carrier_05_CarrierNumber" AT %IW608 : Word;   // CARRIER NUMBER
   "Carrier_05_G120DControlWord" AT %IW610 : Word;   // G120D_STW1_CONTROL
   "Carrier_05_G120DControlWord.0" AT %I610.0 : Bool;   // Bit_00_ON
   "Carrier_05_G120DControlWord.1" AT %I610.1 : Bool;   // Bit_01_AUS2_INH
   "Carrier_05_G120DControlWord.2" AT %I610.2 : Bool;   // Bit_02_AUS3_STOP
   "Carrier_05_G120DControlWord.3" AT %I610.3 : Bool;   // Bit_03_EN
   "Carrier_05_G120DControlWord.4" AT %I610.4 : Bool;   // Bit_04_EN_RAMP
   "Carrier_05_G120DControlWord.5" AT %I610.5 : Bool;   // Bit_05_START_RAMP
   "Carrier_05_G120DControlWord.6" AT %I610.6 : Bool;   // Bit_06_SETPOINT
   "Carrier_05_G120DControlWord.7" AT %I610.7 : Bool;   // Bit_07_RESET
   "Carrier_05_G120DControlWord.8" AT %I611.0 : Bool;   // Bit_08_JOG_R
   "Carrier_05_G120DControlWord.9" AT %I611.1 : Bool;   // Bit_09_JOG_L
   "Carrier_05_G120DControlWord.10" AT %I611.2 : Bool;   // Bit_10_CONTR_PLC
   "Carrier_05_G120DControlWord.11" AT %I611.3 : Bool;   // Bit_11_REVERSE
   "Carrier_05_G120DControlWord.12" AT %I611.4 : Bool;   // Bit_12_BRAKE_RELEASE
   "Carrier_05_G120DControlWord.13" AT %I611.5 : Bool;   // Bit_13_DDS
   "Carrier_05_G120DControlWord.14" AT %I611.6 : Bool;   // Bit_14_DO0
   "Carrier_05_G120DControlWord.15" AT %I611.7 : Bool;   // Bit_15_DO1
   "Carrier_05_G120DStatusWord" AT %IW612 : Word;   // G120D_ZSW1_STATUS
   "Carrier_05_G120DStatusWord.0" AT %I612.0 : Bool;   // Bit_00_READY_RUN
   "Carrier_05_G120DStatusWord.1" AT %I612.1 : Bool;   // Bit_01_READY_ON
   "Carrier_05_G120DStatusWord.2" AT %I612.2 : Bool;   // Bit_02_ENABLE
   "Carrier_05_G120DStatusWord.3" AT %I612.3 : Bool;   // Bit_03_FAULT
   "Carrier_05_G120DStatusWord.4" AT %I612.4 : Bool;   // Bit_04_OFF2
   "Carrier_05_G120DStatusWord.5" AT %I612.5 : Bool;   // Bit_05_OFF3
   "Carrier_05_G120DStatusWord.6" AT %I612.6 : Bool;   // Bit_06_LOCK_OUT
   "Carrier_05_G120DStatusWord.7" AT %I612.7 : Bool;   // Bit_07_WARN
   "Carrier_05_G120DStatusWord.8" AT %I613.0 : Bool;   // Bit_08_NO_DEVIATION
   "Carrier_05_G120DStatusWord.9" AT %I613.1 : Bool;   // Bit_09_CONTR_PLC
   "Carrier_05_G120DStatusWord.10" AT %I613.2 : Bool;   // Bit_10_F_MAX
   "Carrier_05_G120DStatusWord.11" AT %I613.3 : Bool;   // Bit_11_LIMIT_REACHED
   "Carrier_05_G120DStatusWord.12" AT %I613.4 : Bool;   // Bit_12_BRAKE_OPEN
   "Carrier_05_G120DStatusWord.13" AT %I613.5 : Bool;   // Bit_13_NO_OVERTEMP
   "Carrier_05_G120DStatusWord.14" AT %I613.6 : Bool;   // Bit_14_CW_CCW
   "Carrier_05_G120DStatusWord.15" AT %I613.7 : Bool;   // Bit_15_OVERL
   "Carrier_05_Slot2_Input" AT %IW614 : Word;   // SLOT 2 INPUT WORD
   "Carrier_05_CrashDetectSW" AT %I614.0 : Bool;   // CRASH DETECT SW
   "Carrier_05_SpareSafetyInput(2_1)" AT %I614.1 : Bool;   // SPARE SAFETY INPUT
   "Carrier_05_SpareSafetyInput(2_2)" AT %I614.2 : Bool;   // SPARE SAFETY INPUT
   "Carrier_05_SpareSafetyInput(2_3)" AT %I614.3 : Bool;   // SPARE SAFETY INPUT
   "Carrier_05_SpareSafetyInput(2_4)" AT %I614.4 : Bool;   // SPARE SAFETY INPUT
   "Carrier_05_SpareSafetyInput(2_5)" AT %I614.5 : Bool;   // SPARE SAFETY INPUT
   "Carrier_05_SpareSafetyInput(2_6)" AT %I614.6 : Bool;   // SPARE SAFETY INPUT
   "Carrier_05_SpareSafetyInput(2_7)" AT %I614.7 : Bool;   // SPARE SAFETY INPUT
   "Carrier_05_Slot3_SafetyOutput" AT %IW615 : Word;   // SLOT 3 SAFETY OUTPUT WORD